
screen "0113_SettingShiftPlan" 1280x800, template "Navigation"
   on GenerateScreen: SetTag("Recipe_Appearance_Control", 1); function_b431313b("Shifttime", U 1, N)
   on ClearScreen: function_f38ba6b2("Shifttime", U 1, 1, 0, N)
   Button "Button_1" at 612,704 size 245x55; TextOff 'Next Shift'
   TextField "Text field_8" at 305,167 size 204x48; Text 'Shift 1'
   TextField "Text field_9" at 517,167 size 204x48; Text 'Shift 2'
   TextField "Text field_10" at 729,167 size 204x48; Text 'Shift 3'
   TextField "Text field_11" at 941,167 size 204x48; Text 'Shift 4'
   Button "Button_3" at 326,104 size 451x32; TextOff 'Setting Shift Plan'
   Button "b_ShifProto_ShotCounter_1" at 208,713 size 60x60; TextOff 'Shot Counter'; PictureList "ico_ShiftProtocol"
      Appearance <- "Recipe_Appearance_Control"
      ProcessValue <- "Recipe_Appearance_Control"
   Button "b_Shiftproto_shiftproto" at 208,713 size 60x60; TextOff 'Shift proto'
      Appearance <- "Recipe_Appearance_Control"
      on Click: ActivateScreen("0112_Shift protocol", 0); SetTag("Recipe_Appearance_Control", 2)
   Button "b_SC" at 478,713 size 60x60; TextOff 'Shot Counter'; PictureList "ico_ShotCounter"
      on Press: ActivateScreen("0891_Shotcounter MixingHead", 0); SetTag("Recipe_Appearance_Control", 5)
      Appearance <- "Recipe_Appearance_Control"
      ProcessValue <- "Recipe_Appearance_Control"
   Button "b_SC_1" at 478,713 size 60x60; TextOff 'Shot Counter'
      Appearance <- "Recipe_Appearance_Control"
      on Click: ActivateScreen("0891_Shotcounter MixingHead", 0); SetTag("Recipe_Appearance_Control", 5)
   Button "b_Shift_Plan" at 118,713 size 60x60; TextOff 'Shift Plan'; PictureList "ico_ShiftPlan"
      on Press: ActivateScreen("0113_SettingShiftPlan", 0); SetTag("Recipe_Appearance_Control", 1)
      Appearance <- "Recipe_Appearance_Control"
      ProcessValue <- "Recipe_Appearance_Control"
   Button "b_Shift_Plan_1" at 118,713 size 60x60; TextOff 'Shift Plan'
      Appearance <- "Recipe_Appearance_Control"
      on Click: "SettingShiftPlan"(); ActivateScreen("0113_SettingShiftPlan", 0); SetTag("Recipe_Appearance_Control", 1)
   Button "b_LS_Lastshot" at 298,713 size 60x60; TextOff 'Last Shot'; PictureList "ico_LastShot"
      on Press: ActivateScreen("0036_Last Shot", 0); SetTag("Recipe_Appearance_Control", 3)
      Appearance <- "Recipe_Appearance_Control"
      ProcessValue <- "Recipe_Appearance_Control"
   Button "b_LS_Lastshot_1" at 298,713 size 60x60; TextOff 'Last Shot'
      Appearance <- "Recipe_Appearance_Control"
      on Click: ActivateScreen("0036_Last Shot", 0); SetTag("Recipe_Appearance_Control", 3)
   Button "b_Consumtion" at 388,713 size 60x60; TextOff 'Consumtion / Consum'; PictureList "ico_consum"
      on Press: ActivateScreen("0890_Consumption", 0); SetTag("Recipe_Appearance_Control", 4)
      Appearance <- "Recipe_Appearance_Control"
      ProcessValue <- "Recipe_Appearance_Control"
   Button "b_Consumtion_1" at 388,713 size 60x60; TextOff 'Consumtion / Consum'
      Appearance <- "Recipe_Appearance_Control"
      on Click: ActivateScreen("0890_Consumption", 0); SetTag("Recipe_Appearance_Control", 4)
   TextField "Text field_1" at 134,234 size 152x60; Text 'Monday'
   TextField "Text field_2" at 134,298 size 152x60; Text 'Tuesday'
   TextField "Text field_3" at 134,362 size 152x60; Text 'Wenesday'
   TextField "Text field_4" at 134,426 size 152x60; Text 'Thrusday'
   TextField "Text field_5" at 134,490 size 152x60; Text 'Friday'
   TextField "Text field_6" at 134,554 size 152x60; Text 'Saturday'
   TextField "Text field_7" at 134,618 size 152x60; Text 'Sunday'
   IOField "I/O field_1" at 303,298 size 135x60; Authorization "Operate"; FormatPattern 9999999999999999999999999999999999999999
      on OnFinishInput: "SettingShiftPlan"(); "Shifttime_write"()
      ProcessValue <- "Shift_2_1"
   IOField "I/O field_2" at 303,362 size 135x60; Authorization "Operate"; FormatPattern 9999999999999999999999999999999999999999
      on OnFinishInput: "SettingShiftPlan"(); "Shifttime_write"()
      ProcessValue <- "Shift_3_1"
   IOField "I/O field_3" at 303,426 size 135x60; Authorization "Operate"; FormatPattern 9999999999999999999999999999999999999999
      on OnFinishInput: "SettingShiftPlan"(); "Shifttime_write"()
      ProcessValue <- "Shift_4_1"
   IOField "I/O field_4" at 303,490 size 135x60; Authorization "Operate"; FormatPattern 9999999999999999999999999999999999999999
      on OnFinishInput: "SettingShiftPlan"(); "Shifttime_write"()
      ProcessValue <- "Shift_5_1"
   IOField "I/O field_5" at 303,554 size 135x60; Authorization "Operate"; FormatPattern 9999999999999999999999999999999999999999
      on OnFinishInput: "SettingShiftPlan"(); "Shifttime_write"()
      ProcessValue <- "Shift_6_1"
   IOField "I/O field_6" at 303,618 size 135x60; Authorization "Operate"; FormatPattern 9999999999999999999999999999999999999999
      on OnFinishInput: "SettingShiftPlan"(); "Shifttime_write"()
      ProcessValue <- "Shift_7_1"
   IOField "I/O field_7" at 303,234 size 135x60; Authorization "Operate"; FormatPattern 9999999999999999999999999999999999999999
      on OnFinishInput: "SettingShiftPlan"(); "Shifttime_write"()
      ProcessValue <- "Shift_1_1"
   IOField "I/O field_8" at 515,298 size 135x60; Authorization "Operate"; FormatPattern 9999999999999999999999999999999999999999
      on OnFinishInput: "SettingShiftPlan"(); "Shifttime_write"()
      ProcessValue <- "Shift_2_2"
   IOField "I/O field_9" at 515,362 size 135x60; Authorization "Operate"; FormatPattern 9999999999999999999999999999999999999999
      on OnFinishInput: "SettingShiftPlan"(); "Shifttime_write"()
      ProcessValue <- "Shift_3_2"
   IOField "I/O field_10" at 515,426 size 135x60; Authorization "Operate"; FormatPattern 9999999999999999999999999999999999999999
      on OnFinishInput: "SettingShiftPlan"(); "Shifttime_write"()
      ProcessValue <- "Shift_4_2"
   IOField "I/O field_11" at 515,490 size 135x60; Authorization "Operate"; FormatPattern 9999999999999999999999999999999999999999
      on OnFinishInput: "SettingShiftPlan"(); "Shifttime_write"()
      ProcessValue <- "Shift_5_2"
   IOField "I/O field_12" at 515,554 size 135x60; Authorization "Operate"; FormatPattern 9999999999999999999999999999999999999999
      on OnFinishInput: "SettingShiftPlan"(); "Shifttime_write"()
      ProcessValue <- "Shift_6_2"
   IOField "I/O field_13" at 515,618 size 135x60; Authorization "Operate"; FormatPattern 9999999999999999999999999999999999999999
      on OnFinishInput: "SettingShiftPlan"(); "Shifttime_write"()
      ProcessValue <- "Shift_7_2"
   IOField "I/O field_14" at 515,234 size 135x60; Authorization "Operate"; FormatPattern 9999999999999999999999999999999999999999
      on OnFinishInput: "SettingShiftPlan"(); "Shifttime_write"()
      ProcessValue <- "Shift_1_2"
   IOField "I/O field_15" at 727,298 size 135x60; Authorization "Operate"; FormatPattern 9999999999999999999999999999999999999999
      on OnFinishInput: "SettingShiftPlan"(); "Shifttime_write"()
      ProcessValue <- "Shift_2_3"
   IOField "I/O field_16" at 727,362 size 135x60; Authorization "Operate"; FormatPattern 9999999999999999999999999999999999999999
      on OnFinishInput: "SettingShiftPlan"(); "Shifttime_write"()
      ProcessValue <- "Shift_3_3"
   IOField "I/O field_17" at 727,426 size 135x60; Authorization "Operate"; FormatPattern 9999999999999999999999999999999999999999
      on OnFinishInput: "SettingShiftPlan"(); "Shifttime_write"()
      ProcessValue <- "Shift_4_3"
   IOField "I/O field_18" at 727,490 size 135x60; Authorization "Operate"; FormatPattern 9999999999999999999999999999999999999999
      on OnFinishInput: "SettingShiftPlan"(); "Shifttime_write"()
      ProcessValue <- "Shift_5_3"
   IOField "I/O field_19" at 727,554 size 135x60; Authorization "Operate"; FormatPattern 9999999999999999999999999999999999999999
      on OnFinishInput: "SettingShiftPlan"(); "Shifttime_write"()
      ProcessValue <- "Shift_6_3"
   IOField "I/O field_20" at 727,618 size 135x60; Authorization "Operate"; FormatPattern 9999999999999999999999999999999999999999
      on OnFinishInput: "SettingShiftPlan"(); "Shifttime_write"()
      ProcessValue <- "Shift_7_3"
   IOField "I/O field_21" at 727,234 size 135x60; Authorization "Operate"; FormatPattern 9999999999999999999999999999999999999999
      on OnFinishInput: "SettingShiftPlan"(); "Shifttime_write"()
      ProcessValue <- "Shift_1_3"
   IOField "I/O field_23" at 939,298 size 135x60; Authorization "Operate"; FormatPattern 9999999999999999999999999999999999999999
      on OnFinishInput: "SettingShiftPlan"(); "Shifttime_write"()
      ProcessValue <- "Shift_2_4"
   IOField "I/O field_24" at 939,362 size 135x60; Authorization "Operate"; FormatPattern 9999999999999999999999999999999999999999
      on OnFinishInput: "SettingShiftPlan"(); "Shifttime_write"()
      ProcessValue <- "Shift_3_4"
   IOField "I/O field_25" at 939,426 size 135x60; Authorization "Operate"; FormatPattern 9999999999999999999999999999999999999999
      on OnFinishInput: "SettingShiftPlan"(); "Shifttime_write"()
      ProcessValue <- "Shift_4_4"
   IOField "I/O field_26" at 939,490 size 135x60; Authorization "Operate"; FormatPattern 9999999999999999999999999999999999999999
      on OnFinishInput: "SettingShiftPlan"(); "Shifttime_write"()
      ProcessValue <- "Shift_5_4"
   IOField "I/O field_27" at 939,554 size 135x60; Authorization "Operate"; FormatPattern 9999999999999999999999999999999999999999
      on OnFinishInput: "SettingShiftPlan"(); "Shifttime_write"()
      ProcessValue <- "Shift_6_4"
   IOField "I/O field_28" at 939,618 size 135x60; Authorization "Operate"; FormatPattern 9999999999999999999999999999999999999999
      on OnFinishInput: "SettingShiftPlan"(); "Shifttime_write"()
      ProcessValue <- "Shift_7_4"
   IOField "I/O field_29" at 939,234 size 135x60; Authorization "Operate"; FormatPattern 9999999999999999999999999999999999999999
      on OnFinishInput: "SettingShiftPlan"(); "Shifttime_write"()
      ProcessValue <- "Shift_1_4"
   Button "check_shift1_1" at 446,298 size 61x60; TextOff 'Text'; PictureOff "download"; PictureList "Check_Uncheck"; Authorization "Operate"
      on Click: InvertBit("Shift_En_2_1")
      on Change: "SettingShiftPlan"(); "Shifttime_write"()
      ProcessValue <- "Shift_En_2_1"
   Button "check_shift1_2" at 446,362 size 61x60; TextOff 'Text'; PictureOff "download"; PictureList "Check_Uncheck"; Authorization "Operate"
      on Click: InvertBit("Shift_En_3_1")
      on Change: "SettingShiftPlan"(); "Shifttime_write"()
      ProcessValue <- "Shift_En_3_1"
   Button "check_shift1_3" at 446,426 size 61x60; TextOff 'Text'; PictureOff "download"; PictureList "Check_Uncheck"; Authorization "Operate"
      on Click: InvertBit("Shift_En_4_1")
      on Change: "SettingShiftPlan"(); "Shifttime_write"()
      ProcessValue <- "Shift_En_4_1"
   Button "check_shift1_4" at 446,490 size 61x60; TextOff 'Text'; PictureOff "download"; PictureList "Check_Uncheck"; Authorization "Operate"
      on Click: InvertBit("Shift_En_5_1")
      on Change: "SettingShiftPlan"(); "Shifttime_write"()
      ProcessValue <- "Shift_En_5_1"
   Button "check_shift1_5" at 446,554 size 61x60; TextOff 'Text'; PictureOff "download"; PictureList "Check_Uncheck"; Authorization "Operate"
      on Click: InvertBit("Shift_En_6_1")
      on Change: "SettingShiftPlan"(); "Shifttime_write"()
      ProcessValue <- "Shift_En_6_1"
   Button "check_shift1_6" at 446,618 size 61x60; TextOff 'Text'; PictureOff "download"; PictureList "Check_Uncheck"; Authorization "Operate"
      on Click: InvertBit("Shift_En_7_1")
      on Change: "SettingShiftPlan"(); "Shifttime_write"()
      ProcessValue <- "Shift_En_7_1"
   Button "check_shift1_7" at 446,234 size 61x60; TextOff 'Text'; PictureOff "download"; PictureList "Check_Uncheck"; Authorization "Operate"
      on Click: InvertBit("Shift_En_1_1")
      on Change: "SettingShiftPlan"(); "Shifttime_write"()
      ProcessValue <- "Shift_En_1_1"
   Button "check_shift4_1" at 1084,298 size 61x60; TextOff 'Text'; PictureOff "download"; PictureList "Check_Uncheck"; Authorization "Operate"
      on Click: InvertBit("Shift_En_2_4")
      on Change: "SettingShiftPlan"(); "Shifttime_write"()
      ProcessValue <- "Shift_En_2_4"
   Button "check_shift4_2" at 1084,362 size 61x60; TextOff 'Text'; PictureOff "download"; PictureList "Check_Uncheck"; Authorization "Operate"
      on Click: InvertBit("Shift_En_3_4")
      on Change: "SettingShiftPlan"(); "Shifttime_write"()
      ProcessValue <- "Shift_En_3_4"
   Button "check_shift4_3" at 1084,426 size 61x60; TextOff 'Text'; PictureOff "download"; PictureList "Check_Uncheck"; Authorization "Operate"
      on Click: InvertBit("Shift_En_4_4")
      on Change: "SettingShiftPlan"(); "Shifttime_write"()
      ProcessValue <- "Shift_En_4_4"
   Button "check_shift4_4" at 1084,490 size 61x60; TextOff 'Text'; PictureOff "download"; PictureList "Check_Uncheck"; Authorization "Operate"
      on Click: InvertBit("Shift_En_5_4")
      on Change: "SettingShiftPlan"(); "Shifttime_write"()
      ProcessValue <- "Shift_En_5_4"
   Button "check_shift4_5" at 1084,554 size 61x60; TextOff 'Text'; PictureOff "download"; PictureList "Check_Uncheck"; Authorization "Operate"
      on Click: InvertBit("Shift_En_6_4")
      on Change: "SettingShiftPlan"(); "Shifttime_write"()
      ProcessValue <- "Shift_En_6_4"
   Button "check_shift4_6" at 1084,618 size 61x60; TextOff 'Text'; PictureOff "download"; PictureList "Check_Uncheck"; Authorization "Operate"
      on Click: InvertBit("Shift_En_7_4")
      on Change: "SettingShiftPlan"(); "Shifttime_write"()
      ProcessValue <- "Shift_En_7_4"
   Button "check_shift4_7" at 1084,234 size 61x60; TextOff 'Text'; PictureOff "download"; PictureList "Check_Uncheck"; Authorization "Operate"
      on Click: InvertBit("Shift_En_1_4")
      on Change: "SettingShiftPlan"(); "Shifttime_write"()
      ProcessValue <- "Shift_En_1_4"
   Button "check_shift3_1" at 870,298 size 61x60; TextOff 'Text'; PictureOff "download"; PictureList "Check_Uncheck"; Authorization "Operate"
      on Click: InvertBit("Shift_En_2_3")
      on Change: "SettingShiftPlan"(); "Shifttime_write"()
      ProcessValue <- "Shift_En_2_3"
   Button "check_shift3_2" at 870,362 size 61x60; TextOff 'Text'; PictureOff "download"; PictureList "Check_Uncheck"; Authorization "Operate"
      on Click: InvertBit("Shift_En_3_3")
      on Change: "SettingShiftPlan"(); "Shifttime_write"()
      ProcessValue <- "Shift_En_3_3"
   Button "check_shift3_3" at 870,426 size 61x60; TextOff 'Text'; PictureOff "download"; PictureList "Check_Uncheck"; Authorization "Operate"
      on Click: InvertBit("Shift_En_4_3")
      on Change: "SettingShiftPlan"(); "Shifttime_write"()
      ProcessValue <- "Shift_En_4_3"
   Button "check_shift3_4" at 870,490 size 61x60; TextOff 'Text'; PictureOff "download"; PictureList "Check_Uncheck"; Authorization "Operate"
      on Click: InvertBit("Shift_En_5_3")
      on Change: "SettingShiftPlan"(); "Shifttime_write"()
      ProcessValue <- "Shift_En_5_3"
   Button "check_shift3_5" at 870,554 size 61x60; TextOff 'Text'; PictureOff "download"; PictureList "Check_Uncheck"; Authorization "Operate"
      on Click: InvertBit("Shift_En_6_3")
      on Change: "SettingShiftPlan"(); "Shifttime_write"()
      ProcessValue <- "Shift_En_6_3"
   Button "check_shift3_6" at 870,618 size 61x60; TextOff 'Text'; PictureOff "download"; PictureList "Check_Uncheck"; Authorization "Operate"
      on Click: InvertBit("Shift_En_7_3")
      on Change: "SettingShiftPlan"(); "Shifttime_write"()
      ProcessValue <- "Shift_En_7_3"
   Button "check_shift3_7" at 870,234 size 61x60; TextOff 'Text'; PictureOff "download"; PictureList "Check_Uncheck"; Authorization "Operate"
      on Click: InvertBit("Shift_En_1_3")
      on Change: "SettingShiftPlan"(); "Shifttime_write"()
      ProcessValue <- "Shift_En_1_3"
   Button "check_shift2_1" at 659,298 size 61x60; TextOff 'Text'; PictureOff "download"; PictureList "Check_Uncheck"; Authorization "Operate"
      on Click: InvertBit("Shift_En_2_2")
      on Change: "SettingShiftPlan"(); "Shifttime_write"()
      ProcessValue <- "Shift_En_2_2"
   Button "check_shift2_2" at 659,362 size 61x60; TextOff 'Text'; PictureOff "download"; PictureList "Check_Uncheck"; Authorization "Operate"
      on Click: InvertBit("Shift_En_3_2")
      on Change: "SettingShiftPlan"(); "Shifttime_write"()
      ProcessValue <- "Shift_En_3_2"
   Button "check_shift2_3" at 659,426 size 61x60; TextOff 'Text'; PictureOff "download"; PictureList "Check_Uncheck"; Authorization "Operate"
      on Click: InvertBit("Shift_En_4_2")
      on Change: "SettingShiftPlan"(); "Shifttime_write"()
      ProcessValue <- "Shift_En_4_2"
   Button "check_shift2_4" at 659,490 size 61x60; TextOff 'Text'; PictureOff "download"; PictureList "Check_Uncheck"; Authorization "Operate"
      on Click: InvertBit("Shift_En_5_2")
      on Change: "SettingShiftPlan"(); "Shifttime_write"()
      ProcessValue <- "Shift_En_5_2"
   Button "check_shift2_5" at 659,554 size 61x60; TextOff 'Text'; PictureOff "download"; PictureList "Check_Uncheck"; Authorization "Operate"
      on Click: InvertBit("Shift_En_6_2")
      on Change: "SettingShiftPlan"(); "Shifttime_write"()
      ProcessValue <- "Shift_En_6_2"
   Button "check_shift2_6" at 659,618 size 61x60; TextOff 'Text'; PictureOff "download"; PictureList "Check_Uncheck"; Authorization "Operate"
      on Click: InvertBit("Shift_En_7_2")
      on Change: "SettingShiftPlan"(); "Shifttime_write"()
      ProcessValue <- "Shift_En_7_2"
   Button "check_shift2_7" at 659,234 size 61x60; TextOff 'Text'; PictureOff "download"; PictureList "Check_Uncheck"; Authorization "Operate"
      on Click: InvertBit("Shift_En_1_2")
      on Change: "SettingShiftPlan"(); "Shifttime_write"()
      ProcessValue <- "Shift_En_1_2"
   IOField "I/O field_30" at 894,704 size 227x55; FormatPattern 9999999999999999999999999999999999999999
      ProcessValue <- "Next shift"

screen "0112_Shift protocol" 1280x800, template "Navigation"
   on GenerateScreen: SetTag("Recipe_Appearance_Control", 2); function_b431313b("ShiftProtocol", U 1, N)
   on ClearScreen: SetTag("Recipe_Appearance_Control", 0)
   TextField "Text field_1" at 109,205 size 57x47; Text '1.'
   TextField "Text field_2" at 109,270 size 57x47; Text '2.'
   TextField "Text field_3" at 109,335 size 57x47; Text '3.'
   TextField "Text field_4" at 109,402 size 57x47; Text '4.'
   TextField "Text field_5" at 109,469 size 57x47; Text '5.'
   TextField "Text field_6" at 109,537 size 57x47; Text '6.'
   TextField "Text field_7" at 109,605 size 57x47; Text '7.'
   IOField "shiftproto_1" at 176,205 size 267x47; FormatPattern 9999999999999999999999999999999999999999
      ProcessValue <- "Shift_Protocol_1"
   IOField "I/O field_2" at 176,270 size 267x47; FormatPattern 9999999999999999999999999999999999999999
      ProcessValue <- "Shift_Protocol_2"
   IOField "I/O field_3" at 176,335 size 267x47; FormatPattern 9999999999999999999999999999999999999999
      ProcessValue <- "Shift_Protocol_3"
   IOField "I/O field_4" at 176,402 size 267x47; FormatPattern 9999999999999999999999999999999999999999
      ProcessValue <- "Shift_Protocol_4"
   IOField "I/O field_5" at 176,469 size 267x47; FormatPattern 9999999999999999999999999999999999999999
      ProcessValue <- "Shift_Protocol_5"
   IOField "I/O field_6" at 176,537 size 267x47; FormatPattern 9999999999999999999999999999999999999999
      ProcessValue <- "Shift_Protocol_6"
   IOField "I/O field_7" at 176,605 size 267x47; FormatPattern 9999999999999999999999999999999999999999
      ProcessValue <- "Shift_Protocol_7"
   IOField "I/O field_8" at 543,205 size 267x47; FormatPattern 9999999999999999999999999999999999999999
      ProcessValue <- "Shift_Protocol_8"
   IOField "I/O field_9" at 902,205 size 267x47; FormatPattern 9999999999999999999999999999999999999999
      ProcessValue <- "Shift_Protocol_15"
   IOField "I/O field_10" at 543,270 size 267x47; FormatPattern 9999999999999999999999999999999999999999
      ProcessValue <- "Shift_Protocol_9"
   IOField "I/O field_11" at 543,335 size 267x47; FormatPattern 9999999999999999999999999999999999999999
      ProcessValue <- "Shift_Protocol_10"
   IOField "I/O field_12" at 543,402 size 267x47; FormatPattern 9999999999999999999999999999999999999999
      ProcessValue <- "Shift_Protocol_11"
   IOField "I/O field_13" at 543,469 size 267x47; FormatPattern 9999999999999999999999999999999999999999
      ProcessValue <- "Shift_Protocol_12"
   IOField "I/O field_14" at 543,537 size 267x47; FormatPattern 9999999999999999999999999999999999999999
      ProcessValue <- "Shift_Protocol_13"
   IOField "I/O field_15" at 543,605 size 267x47; FormatPattern 9999999999999999999999999999999999999999
      ProcessValue <- "Shift_Protocol_14"
   IOField "I/O field_16" at 902,270 size 267x47; FormatPattern 9999999999999999999999999999999999999999
      ProcessValue <- "Shift_Protocol_16"
   IOField "I/O field_17" at 902,335 size 267x47; FormatPattern 9999999999999999999999999999999999999999
      ProcessValue <- "Shift_Protocol_17"
   IOField "I/O field_18" at 902,402 size 267x47; FormatPattern 9999999999999999999999999999999999999999
      ProcessValue <- "Shift_Protocol_18"
   IOField "I/O field_19" at 902,469 size 267x47; FormatPattern 9999999999999999999999999999999999999999
      ProcessValue <- "Shift_Protocol_19"
   IOField "I/O field_20" at 902,537 size 267x47; FormatPattern 9999999999999999999999999999999999999999
      ProcessValue <- "Shift_Protocol_20"
   IOField "I/O field_21" at 902,605 size 267x47; FormatPattern 9999999999999999999999999999999999999999
      ProcessValue <- "Shift_Protocol_21"
   TextField "Text field_8" at 474,205 size 57x47; Text '8.'
   TextField "Text field_9" at 474,270 size 57x47; Text '9.'
   TextField "Text field_10" at 474,335 size 57x47; Text '10.'
   TextField "Text field_11" at 474,402 size 57x47; Text '11.'
   TextField "Text field_12" at 474,469 size 57x47; Text '12.'
   TextField "Text field_13" at 474,537 size 57x47; Text '13.'
   TextField "Text field_14" at 474,605 size 57x47; Text '14.'
   TextField "Text field_15" at 836,205 size 57x47; Text '15.'
   TextField "Text field_16" at 836,270 size 57x47; Text '16.'
   TextField "Text field_17" at 836,335 size 57x47; Text '17.'
   TextField "Text field_18" at 836,402 size 57x47; Text '18.'
   TextField "Text field_19" at 836,469 size 57x47; Text '19.'
   TextField "Text field_20" at 836,537 size 57x47; Text '20.'
   TextField "Text field_21" at 836,605 size 57x47; Text '21.'
   Button "Button_3" at 326,104 size 451x32; TextOff 'Shift Protocol'
   Button "b_spare" at 1000,713 size 60x60; TextOff 'Text'; PictureOff "USB_1"
      on Click: function_ea909784("ShiftProtocol", U 0, '\Storage Card USB\record.csv', 1, 1, N)
   Button "Button_1" at 172,202 size 276x54; TextOff 'Text'
      on Click: SetTag("Archive Alarm Number", 1); SetTag("Archived Alarm Control", 1); "CopyAlarmLogView"(); ActivateScreen("0013_Archive Alarm", 0)
   Button "b_ShifProto_ShotCounter_1" at 208,713 size 60x60; TextOff 'Shot Counter'; PictureList "ico_ShiftProtocol"
      ProcessValue <- "Recipe_Appearance_Control"
      Appearance <- "Recipe_Appearance_Control"
   Button "b_Shiftproto_shiftproto" at 208,713 size 60x60; TextOff 'Shift proto'
      on Click: ActivateScreen("0112_Shift protocol", 0); SetTag("Recipe_Appearance_Control", 2)
      Appearance <- "Recipe_Appearance_Control"
   Button "b_SC" at 478,713 size 60x60; TextOff 'Shot Counter'; PictureList "ico_ShotCounter"
      on Press: ActivateScreen("0891_Shotcounter MixingHead", 0); SetTag("Recipe_Appearance_Control", 5)
      Appearance <- "Recipe_Appearance_Control"
      ProcessValue <- "Recipe_Appearance_Control"
   Button "b_SC_1" at 478,713 size 60x60; TextOff 'Shot Counter'
      on Click: ActivateScreen("0891_Shotcounter MixingHead", 0); SetTag("Recipe_Appearance_Control", 5)
      Appearance <- "Recipe_Appearance_Control"
   Button "b_Shift_Plan" at 118,713 size 60x60; TextOff 'Shift Plan'; PictureList "ico_ShiftPlan"
      on Press: ActivateScreen("0113_SettingShiftPlan", 0); SetTag("Recipe_Appearance_Control", 1)
      Appearance <- "Recipe_Appearance_Control"
      ProcessValue <- "Recipe_Appearance_Control"
   Button "b_Shift_Plan_1" at 118,713 size 60x60; TextOff 'Shift Plan'
      on Click: "SettingShiftPlan"(); ActivateScreen("0113_SettingShiftPlan", 0); SetTag("Recipe_Appearance_Control", 1)
      Appearance <- "Recipe_Appearance_Control"
   Button "b_LS_Lastshot" at 298,713 size 60x60; TextOff 'Last Shot'; PictureList "ico_LastShot"
      on Press: ActivateScreen("0036_Last Shot", 0); SetTag("Recipe_Appearance_Control", 3)
      Appearance <- "Recipe_Appearance_Control"
      ProcessValue <- "Recipe_Appearance_Control"
   Button "b_LS_Lastshot_1" at 298,713 size 60x60; TextOff 'Last Shot'
      on Click: ActivateScreen("0036_Last Shot", 0); SetTag("Recipe_Appearance_Control", 3)
      Appearance <- "Recipe_Appearance_Control"
   Button "b_Consumtion" at 388,713 size 60x60; TextOff 'Consumtion / Consum'; PictureList "ico_consum"
      on Press: ActivateScreen("0890_Consumption", 0); SetTag("Recipe_Appearance_Control", 4)
      Appearance <- "Recipe_Appearance_Control"
      ProcessValue <- "Recipe_Appearance_Control"
   Button "b_Consumtion_1" at 388,713 size 60x60; TextOff 'Consumtion / Consum'
      on Click: ActivateScreen("0890_Consumption", 0); SetTag("Recipe_Appearance_Control", 4)
      Appearance <- "Recipe_Appearance_Control"
   Button "Button_2" at 172,267 size 276x54; TextOff 'Text'
      on Click: SetTag("Archive Alarm Number", 2); SetTag("Archived Alarm Control", 1); "CopyAlarmLogView"(); ActivateScreen("0013_Archive Alarm", 0)
   Button "Button_4" at 172,332 size 276x54; TextOff 'Text'
      on Click: SetTag("Archive Alarm Number", 3); SetTag("Archived Alarm Control", 1); "CopyAlarmLogView"(); ActivateScreen("0013_Archive Alarm", 0)
   Button "Button_5" at 172,397 size 276x54; TextOff 'Text'
      on Click: SetTag("Archive Alarm Number", 4); SetTag("Archived Alarm Control", 1); "CopyAlarmLogView"(); ActivateScreen("0013_Archive Alarm", 0)
   Button "Button_6" at 172,465 size 276x54; TextOff 'Text'
      on Click: SetTag("Archive Alarm Number", 5); SetTag("Archived Alarm Control", 1); "CopyAlarmLogView"(); ActivateScreen("0013_Archive Alarm", 0)
   Button "Button_7" at 172,535 size 276x54; TextOff 'Text'
      on Click: SetTag("Archive Alarm Number", 6); SetTag("Archived Alarm Control", 1); "CopyAlarmLogView"(); ActivateScreen("0013_Archive Alarm", 0)
   Button "Button_8" at 172,602 size 276x54; TextOff 'Text'
      on Click: SetTag("Archive Alarm Number", 7); SetTag("Archived Alarm Control", 1); "CopyAlarmLogView"(); ActivateScreen("0013_Archive Alarm", 0)
   Button "Button_9" at 540,202 size 276x54; TextOff 'Text'
      on Click: SetTag("Archive Alarm Number", 8); SetTag("Archived Alarm Control", 1); "CopyAlarmLogView"(); ActivateScreen("0013_Archive Alarm", 0)
   Button "Button_10" at 540,267 size 276x54; TextOff 'Text'
      on Click: SetTag("Archive Alarm Number", 9); SetTag("Archived Alarm Control", 1); "CopyAlarmLogView"(); ActivateScreen("0013_Archive Alarm", 0)
   Button "Button_11" at 540,332 size 276x54; TextOff 'Text'
      on Click: SetTag("Archive Alarm Number", 10); SetTag("Archived Alarm Control", 1); "CopyAlarmLogView"(); ActivateScreen("0013_Archive Alarm", 0)
   Button "Button_12" at 540,397 size 276x54; TextOff 'Text'
      on Click: SetTag("Archive Alarm Number", 11); SetTag("Archived Alarm Control", 1); "CopyAlarmLogView"(); ActivateScreen("0013_Archive Alarm", 0)
   Button "Button_13" at 540,465 size 276x54; TextOff 'Text'
      on Click: SetTag("Archive Alarm Number", 12); SetTag("Archived Alarm Control", 1); "CopyAlarmLogView"(); ActivateScreen("0013_Archive Alarm", 0)
   Button "Button_14" at 540,535 size 276x54; TextOff 'Text'
      on Click: SetTag("Archive Alarm Number", 13); SetTag("Archived Alarm Control", 1); "CopyAlarmLogView"(); ActivateScreen("0013_Archive Alarm", 0)
   Button "Button_15" at 540,602 size 276x54; TextOff 'Text'
      on Click: SetTag("Archive Alarm Number", 14); SetTag("Archived Alarm Control", 1); "CopyAlarmLogView"(); ActivateScreen("0013_Archive Alarm", 0)
   Button "Button_16" at 900,202 size 276x54; TextOff 'Text'
      on Click: SetTag("Archive Alarm Number", 15); SetTag("Archived Alarm Control", 1); "CopyAlarmLogView"(); ActivateScreen("0013_Archive Alarm", 0)
   Button "Button_17" at 900,267 size 276x54; TextOff 'Text'
      on Click: SetTag("Archive Alarm Number", 16); SetTag("Archived Alarm Control", 1); "CopyAlarmLogView"(); ActivateScreen("0013_Archive Alarm", 0)
   Button "Button_18" at 900,332 size 276x54; TextOff 'Text'
      on Click: SetTag("Archive Alarm Number", 17); SetTag("Archived Alarm Control", 1); "CopyAlarmLogView"(); ActivateScreen("0013_Archive Alarm", 0)
   Button "Button_19" at 900,397 size 276x54; TextOff 'Text'
      on Click: SetTag("Archive Alarm Number", 18); SetTag("Archived Alarm Control", 1); "CopyAlarmLogView"(); ActivateScreen("0013_Archive Alarm", 0)
   Button "Button_20" at 900,465 size 276x54; TextOff 'Text'
      on Click: SetTag("Archive Alarm Number", 19); SetTag("Archived Alarm Control", 1); "CopyAlarmLogView"(); ActivateScreen("0013_Archive Alarm", 0)
   Button "Button_21" at 900,535 size 276x54; TextOff 'Text'
      on Click: SetTag("Archive Alarm Number", 20); SetTag("Archived Alarm Control", 1); "CopyAlarmLogView"(); ActivateScreen("0013_Archive Alarm", 0)
   Button "Button_22" at 900,602 size 276x54; TextOff 'Text'
      on Click: SetTag("Archive Alarm Number", 21); SetTag("Archived Alarm Control", 1); "CopyAlarmLogView"(); ActivateScreen("0013_Archive Alarm", 0)

screen "0036_Last Shot" 1280x800, template "Navigation"
   on GenerateScreen: SetTag("Recipe_Appearance_Control", 3)
   IOField "Prg_1" at 156,204 size 45x30; FormatPattern 99
      ProcessValue <- "DB918_ShotResultlast10_FilteredShot{1}_StationNo"
   IOField "I/O field_2" at 156,290 size 45x30; FormatPattern 99
      ProcessValue <- "DB918_ShotResultlast10_FilteredShot{2}_StationNo"
   IOField "I/O field_3" at 156,378 size 45x30; FormatPattern 99
      ProcessValue <- "DB918_ShotResultlast10_FilteredShot{3}_StationNo"
   IOField "I/O field_4" at 156,466 size 45x30; FormatPattern 99
      ProcessValue <- "DB918_ShotResultlast10_FilteredShot{4}_StationNo"
   IOField "I/O field_5" at 156,551 size 45x30; FormatPattern 99
      ProcessValue <- "DB918_ShotResultlast10_FilteredShot{5}_StationNo"
   IOField "I/O field_6" at 156,637 size 45x30; FormatPattern 99
      ProcessValue <- "DB918_ShotResultlast10_FilteredShot{6}_StationNo"
   IOField "I/O field_7" at 209,204 size 45x30; FormatPattern 99
      ProcessValue <- "DB918_ShotResultlast10_FilteredShot{1}_MHNo"
   IOField "I/O field_8" at 209,290 size 45x30; FormatPattern 99
      ProcessValue <- "DB918_ShotResultlast10_FilteredShot{2}_MHNo"
   IOField "I/O field_9" at 209,378 size 45x30; FormatPattern 99
      ProcessValue <- "DB918_ShotResultlast10_FilteredShot{3}_MHNo"
   IOField "I/O field_10" at 209,466 size 45x30; FormatPattern 99
      ProcessValue <- "DB918_ShotResultlast10_FilteredShot{4}_MHNo"
   IOField "I/O field_11" at 209,551 size 45x30; FormatPattern 99
      ProcessValue <- "DB918_ShotResultlast10_FilteredShot{5}_MHNo"
   IOField "I/O field_12" at 209,637 size 45x30; FormatPattern 99
      ProcessValue <- "DB918_ShotResultlast10_FilteredShot{6}_MHNo"
   IOField "I/O field_13" at 262,204 size 45x30; FormatPattern 99
      ProcessValue <- "DB918_ShotResultlast10_FilteredShot{1}_PartNo"
   IOField "I/O field_14" at 262,290 size 45x30; FormatPattern 99
      ProcessValue <- "DB918_ShotResultlast10_FilteredShot{2}_PartNo"
   IOField "I/O field_15" at 262,378 size 45x30; FormatPattern 99
      ProcessValue <- "DB918_ShotResultlast10_FilteredShot{3}_PartNo"
   IOField "I/O field_16" at 262,466 size 45x30; FormatPattern 99
      ProcessValue <- "DB918_ShotResultlast10_FilteredShot{4}_PartNo"
   IOField "I/O field_17" at 262,551 size 45x30; FormatPattern 99
      ProcessValue <- "DB918_ShotResultlast10_FilteredShot{5}_PartNo"
   IOField "I/O field_18" at 262,637 size 45x30; FormatPattern 99
      ProcessValue <- "DB918_ShotResultlast10_FilteredShot{6}_PartNo"
   IOField "I/O field_19" at 314,204 size 102x30; FormatPattern 9999.999
      ProcessValue <- "DB918_ShotResultlast10_FilteredShot{1}_FoamingTime"
   IOField "I/O field_20" at 314,290 size 102x30; FormatPattern 9999.999
      ProcessValue <- "DB918_ShotResultlast10_FilteredShot{2}_FoamingTime"
   IOField "I/O field_21" at 314,378 size 102x30; FormatPattern 9999.999
      ProcessValue <- "DB918_ShotResultlast10_FilteredShot{3}_FoamingTime"
   IOField "I/O field_22" at 314,466 size 102x30; FormatPattern 9999.999
      ProcessValue <- "DB918_ShotResultlast10_FilteredShot{4}_FoamingTime"
   IOField "I/O field_23" at 314,551 size 102x30; FormatPattern 9999.999
      ProcessValue <- "DB918_ShotResultlast10_FilteredShot{5}_FoamingTime"
   IOField "I/O field_24" at 314,637 size 102x30; FormatPattern 9999.999
      ProcessValue <- "DB918_ShotResultlast10_FilteredShot{6}_FoamingTime"
   IOField "I/O field_25" at 422,204 size 102x30; FormatPattern 999999.99
      ProcessValue <- "DB918_ShotResultlast10_FilteredShot{1}_PartWeight"
   IOField "I/O field_26" at 422,290 size 102x30; FormatPattern 999999.99
      ProcessValue <- "DB918_ShotResultlast10_FilteredShot{2}_PartWeight"
   IOField "I/O field_27" at 422,378 size 102x30; FormatPattern 999999.99
      ProcessValue <- "DB918_ShotResultlast10_FilteredShot{3}_PartWeight"
   IOField "I/O field_28" at 422,466 size 102x30; FormatPattern 999999.99
      ProcessValue <- "DB918_ShotResultlast10_FilteredShot{4}_PartWeight"
   IOField "I/O field_29" at 422,551 size 102x30; FormatPattern 999999.99
      ProcessValue <- "DB918_ShotResultlast10_FilteredShot{5}_PartWeight"
   IOField "I/O field_30" at 422,637 size 102x30; FormatPattern 999999.99
      ProcessValue <- "DB918_ShotResultlast10_FilteredShot{6}_PartWeight"
   IOField "I/O field_31" at 717,204 size 102x30; FormatPattern 999999.99
      ProcessValue <- "DB918_ShotResultlast10_FilteredShot{1}_Flow{1}"
   IOField "I/O field_32" at 717,240 size 102x30; FormatPattern 999999.99
      ProcessValue <- "DB918_ShotResultlast10_FilteredShot{1}_Flow{2}"
   IOField "I/O field_33" at 717,290 size 102x30; FormatPattern 999999.99
      ProcessValue <- "DB918_ShotResultlast10_FilteredShot{2}_Flow{1}"
   IOField "I/O field_34" at 717,327 size 102x30; FormatPattern 999999.99
      ProcessValue <- "DB918_ShotResultlast10_FilteredShot{2}_Flow{2}(1)"
   IOField "I/O field_35" at 717,379 size 102x30; FormatPattern 999999.99
      ProcessValue <- "DB918_ShotResultlast10_FilteredShot{3}_Flow{1}"
   IOField "I/O field_36" at 717,413 size 102x30; FormatPattern 999999.99
      ProcessValue <- "DB918_ShotResultlast10_FilteredShot{3}_Flow{2}"
   IOField "I/O field_37" at 717,466 size 102x30; FormatPattern 999999.99
      ProcessValue <- "DB918_ShotResultlast10_FilteredShot{4}_Flow{1}"
   IOField "I/O field_38" at 717,501 size 102x30; FormatPattern 999999.99
      ProcessValue <- "DB918_ShotResultlast10_FilteredShot{4}_Flow{2}"
   IOField "I/O field_39" at 717,551 size 102x30; FormatPattern 999999.99
      ProcessValue <- "DB918_ShotResultlast10_FilteredShot{5}_Flow{1}"
   IOField "I/O field_40" at 717,586 size 102x30; FormatPattern 999999.99
      ProcessValue <- "DB918_ShotResultlast10_FilteredShot{5}_Flow{2}"
   IOField "I/O field_41" at 717,637 size 102x30; FormatPattern 999999.99
      ProcessValue <- "DB918_ShotResultlast10_FilteredShot{6}_Flow{1}"
   IOField "I/O field_42" at 824,204 size 82x30; FormatPattern 999999.99
      ProcessValue <- "DB918_ShotResultlast10_FilteredShot{1}_Pressure{1}"
   IOField "I/O field_43" at 824,240 size 82x30; FormatPattern 999999.99
      ProcessValue <- "DB918_ShotResultlast10_FilteredShot{1}_Pressure{2}"
   IOField "I/O field_44" at 824,290 size 82x30; FormatPattern 999999.99
      ProcessValue <- "DB918_ShotResultlast10_FilteredShot{2}_Pressure{1}"
   IOField "I/O field_45" at 824,327 size 82x30; FormatPattern 999999.99
      ProcessValue <- "DB918_ShotResultlast10_FilteredShot{2}_Pressure{2}"
   IOField "I/O field_46" at 824,378 size 82x30; FormatPattern 999999.99
      ProcessValue <- "DB918_ShotResultlast10_FilteredShot{3}_Pressure{1}"
   IOField "I/O field_47" at 824,413 size 82x30; FormatPattern 999999.99
      ProcessValue <- "DB918_ShotResultlast10_FilteredShot{3}_Pressure{2}"
   IOField "I/O field_48" at 824,466 size 82x30; FormatPattern 999999.99
      ProcessValue <- "DB918_ShotResultlast10_FilteredShot{4}_Pressure{1}"
   IOField "I/O field_49" at 824,501 size 82x30; FormatPattern 999999.99
      ProcessValue <- "DB918_ShotResultlast10_FilteredShot{4}_Pressure{2}"
   IOField "I/O field_50" at 824,551 size 82x30; FormatPattern 999999.99
      ProcessValue <- "DB918_ShotResultlast10_FilteredShot{5}_Pressure{1}"
   IOField "I/O field_51" at 824,586 size 82x30; FormatPattern 999999.99
      ProcessValue <- "DB918_ShotResultlast10_FilteredShot{5}_Pressure{2}"
   IOField "I/O field_52" at 824,637 size 82x30; FormatPattern 999999.99
      ProcessValue <- "DB918_ShotResultlast10_FilteredShot{6}_Pressure{1}"
   IOField "I/O field_53" at 911,204 size 82x30; FormatPattern 999999.99
      ProcessValue <- "DB918_ShotResultlast10_FilteredShot{1}_Mixingratio{1}"
   IOField "I/O field_54" at 911,240 size 82x30; FormatPattern 999999.99
      ProcessValue <- "DB918_ShotResultlast10_FilteredShot{1}_Mixingratio{2}"
   IOField "I/O field_55" at 911,290 size 82x30; FormatPattern 999999.99
      ProcessValue <- "DB918_ShotResultlast10_FilteredShot{2}_Mixingratio{1}"
   IOField "I/O field_56" at 911,327 size 82x30; FormatPattern 999999.99
      ProcessValue <- "DB918_ShotResultlast10_FilteredShot{2}_Mixingratio{2}"
   IOField "I/O field_57" at 911,379 size 82x30; FormatPattern 999999.99
      ProcessValue <- "DB918_ShotResultlast10_FilteredShot{3}_Mixingratio{1}"
   IOField "I/O field_58" at 911,413 size 82x30; FormatPattern 999999.99
      ProcessValue <- "DB918_ShotResultlast10_FilteredShot{3}_Mixingratio{2}"
   IOField "I/O field_59" at 911,466 size 82x30; FormatPattern 999999.99
      ProcessValue <- "DB918_ShotResultlast10_FilteredShot{4}_Mixingratio{1}"
   IOField "I/O field_60" at 911,501 size 82x30; FormatPattern 999999.99
      ProcessValue <- "DB918_ShotResultlast10_FilteredShot{4}_Mixingratio{2}"
   IOField "I/O field_61" at 911,551 size 82x30; FormatPattern 999999.99
      ProcessValue <- "DB918_ShotResultlast10_FilteredShot{5}_Mixingratio{1}"
   IOField "I/O field_62" at 911,586 size 82x30; FormatPattern 999999.99
      ProcessValue <- "DB918_ShotResultlast10_FilteredShot{5}_Mixingratio{2}"
   IOField "I/O field_63" at 911,637 size 82x30; FormatPattern 999999.99
      ProcessValue <- "DB918_ShotResultlast10_FilteredShot{6}_Mixingratio{1}"
   IOField "I/O field_64" at 998,204 size 82x30; FormatPattern 999999.9
      ProcessValue <- "DB918_ShotResultlast10_FilteredShot{1}_Temperature{1}"
   IOField "I/O field_65" at 998,240 size 82x30; FormatPattern 999999.9
      ProcessValue <- "DB918_ShotResultlast10_FilteredShot{1}_Temperature{2}"
   IOField "I/O field_66" at 998,290 size 82x30; FormatPattern 999999.9
      ProcessValue <- "DB918_ShotResultlast10_FilteredShot{2}_Temperature{1}"
   IOField "I/O field_67" at 998,327 size 82x30; FormatPattern 999999.9
      ProcessValue <- "DB918_ShotResultlast10_FilteredShot{2}_Temperature{2}"
   IOField "I/O field_68" at 998,378 size 82x30; FormatPattern 999999.9
      ProcessValue <- "DB918_ShotResultlast10_FilteredShot{3}_Temperature{1}"
   IOField "I/O field_69" at 998,413 size 82x30; FormatPattern 999999.9
      ProcessValue <- "DB918_ShotResultlast10_FilteredShot{3}_Temperature{2}"
   IOField "I/O field_70" at 998,466 size 82x30; FormatPattern 999999.9
      ProcessValue <- "DB918_ShotResultlast10_FilteredShot{4}_Temperature{1}"
   IOField "I/O field_71" at 998,501 size 82x30; FormatPattern 999999.9
      ProcessValue <- "DB918_ShotResultlast10_FilteredShot{4}_Temperature{2}"
   IOField "I/O field_72" at 998,551 size 82x30; FormatPattern 999999.9
      ProcessValue <- "DB918_ShotResultlast10_FilteredShot{5}_Temperature{1}"
   IOField "I/O field_73" at 998,586 size 82x30; FormatPattern 999999.9
      ProcessValue <- "DB918_ShotResultlast10_FilteredShot{5}_Temperature{2}"
   IOField "I/O field_74" at 998,637 size 82x30; FormatPattern 999999.9
      ProcessValue <- "DB918_ShotResultlast10_FilteredShot{6}_Temperature{1}"
   IOField "I/O field_75" at 1085,204 size 82x30; FormatPattern 999999.99
      ProcessValue <- "DB918_ShotResultlast10_FilteredShot{1}_MaterialConsumption{1}"
   IOField "I/O field_76" at 1085,240 size 82x30; FormatPattern 999999.99
      ProcessValue <- "DB918_ShotResultlast10_FilteredShot{1}_MaterialConsumption{2}"
   IOField "I/O field_77" at 1085,290 size 82x30; FormatPattern 999999.99
      ProcessValue <- "DB918_ShotResultlast10_FilteredShot{2}_MaterialConsumption{1}"
   IOField "I/O field_78" at 1085,327 size 82x30; FormatPattern 999999.99
      ProcessValue <- "DB918_ShotResultlast10_FilteredShot{2}_MaterialConsumption{2}"
   IOField "I/O field_79" at 1085,378 size 82x30; FormatPattern 999999.99
      ProcessValue <- "DB918_ShotResultlast10_FilteredShot{3}_MaterialConsumption{1}"
   IOField "I/O field_80" at 1085,413 size 82x30; FormatPattern 999999.99
      ProcessValue <- "DB918_ShotResultlast10_FilteredShot{3}_MaterialConsumption{2}"
   IOField "I/O field_81" at 1085,466 size 82x30; FormatPattern 999999.99
      ProcessValue <- "DB918_ShotResultlast10_FilteredShot{4}_MaterialConsumption{1}"
   IOField "I/O field_82" at 1085,501 size 82x30; FormatPattern 999999.99
      ProcessValue <- "DB918_ShotResultlast10_FilteredShot{4}_MaterialConsumption{2}"
   IOField "I/O field_83" at 1085,551 size 82x30; FormatPattern 999999.99
      ProcessValue <- "DB918_ShotResultlast10_FilteredShot{5}_MaterialConsumption{1}"
   IOField "I/O field_84" at 1085,586 size 82x30; FormatPattern 999999.99
      ProcessValue <- "DB918_ShotResultlast10_FilteredShot{5}_MaterialConsumption{2}"
   IOField "I/O field_85" at 1085,637 size 82x30; FormatPattern 999999.99
      ProcessValue <- "DB918_ShotResultlast10_FilteredShot{6}_MaterialConsumption{1}"
   Button "Button_3" at 326,99 size 451x32; TextOff 'Last Shot'
   IOField "I/O field_86" at 717,674 size 102x30; FormatPattern 999999.99
      ProcessValue <- "DB918_ShotResultlast10_FilteredShot{6}_Flow{2}"
   IOField "I/O field_87" at 824,674 size 82x30; FormatPattern 999999.99
      ProcessValue <- "DB918_ShotResultlast10_FilteredShot{6}_Pressure{2}"
   IOField "I/O field_88" at 911,674 size 82x30; FormatPattern 999999.99
      ProcessValue <- "DB918_ShotResultlast10_FilteredShot{6}_Mixingratio{2}"
   IOField "I/O field_89" at 998,674 size 82x30; FormatPattern 999999.9
      ProcessValue <- "DB918_ShotResultlast10_FilteredShot{6}_Temperature{2}"
   IOField "I/O field_90" at 1085,674 size 82x30; FormatPattern 999999.99
      ProcessValue <- "DB918_ShotResultlast10_FilteredShot{6}_MaterialConsumption{2}"
   Button "Button_14" at 156,145 size 45x33; TextOff 'Prg.'
   Button "Button_15" at 209,145 size 45x33; TextOff 'MH'
   Button "Button_16" at 262,145 size 45x33; TextOff 'PS'
   Button "Button_17" at 314,145 size 102x33; TextOff 'Time'
   Button "Button_18" at 422,145 size 102x33; TextOff 'Weight'
   Button "Button_19" at 530,145 size 182x33; TextOff 'Name'
   Button "Button_20" at 717,145 size 102x33; TextOff 'Flow'
   Button "Button_21" at 825,145 size 82x33; TextOff 'Pressure'
   Button "Button_22" at 912,145 size 82x33; TextOff 'Ratio'
   Button "Button_23" at 998,145 size 82x33; TextOff 'Temp'
   Button "Button_24" at 1085,145 size 82x33; TextOff 'Weight'
   IOField "I/O field_91" at 529,204 size 182x30; FormatPattern ????????????????????
      ProcessValue <- "DB918_ShotResultlast10_FilteredShot{1}_Name{1}"
   IOField "I/O field_92" at 530,240 size 182x30; FormatPattern ????????????????????
      ProcessValue <- "DB918_ShotResultlast10_FilteredShot{1}_Name{2}"
   IOField "I/O field_93" at 530,290 size 182x30; FormatPattern ????????????????????
      ProcessValue <- "DB918_ShotResultlast10_FilteredShot{2}_Name{1}"
   IOField "I/O field_94" at 530,327 size 182x30; FormatPattern ????????????????????
      ProcessValue <- "DB918_ShotResultlast10_FilteredShot{2}_Name{2}"
   IOField "I/O field_95" at 530,378 size 182x30; FormatPattern ????????????????????
      ProcessValue <- "DB918_ShotResultlast10_FilteredShot{3}_Name{1}"
   IOField "I/O field_96" at 530,413 size 182x30; FormatPattern ????????????????????
      ProcessValue <- "DB918_ShotResultlast10_FilteredShot{3}_Name{2}"
   IOField "I/O field_97" at 530,466 size 182x30; FormatPattern ????????????????????
      ProcessValue <- "DB918_ShotResultlast10_FilteredShot{4}_Name{1}"
   IOField "I/O field_98" at 530,501 size 182x30; FormatPattern ????????????????????
      ProcessValue <- "DB918_ShotResultlast10_FilteredShot{4}_Name{2}"
   IOField "I/O field_99" at 530,551 size 182x30; FormatPattern ????????????????????
      ProcessValue <- "DB918_ShotResultlast10_FilteredShot{5}_Name{1}"
   IOField "I/O field_100" at 530,586 size 182x30; FormatPattern ????????????????????
      ProcessValue <- "DB918_ShotResultlast10_FilteredShot{5}_Name{2}"
   IOField "I/O field_101" at 530,637 size 182x30; FormatPattern ????????????????????
      ProcessValue <- "DB918_ShotResultlast10_FilteredShot{6}_Name{1}"
   IOField "I/O field_102" at 530,674 size 182x30; FormatPattern ????????????????????
      ProcessValue <- "DB918_ShotResultlast10_FilteredShot{6}_Name{2}"
   GraphicView "Graphic view_1" at 104,204 size 45x30; Picture "cp2"
      Visibility <- "DB918_ShotResultlast10_FilteredShot{1}_PartShotDisableService"
   GraphicView "Graphic view_2" at 104,204 size 45x30; Picture "manual mode"
      Visibility <- "DB918_ShotResultlast10_FilteredShot{1}_StatusBitManualShot"
   GraphicView "Graphic view_3" at 104,204 size 45x30; Picture "automatic mode"
      Visibility <- "DB918_ShotResultlast10_FilteredShot{1}_StatusBitAutomaticShot"
   GraphicView "Graphic view_4" at 104,290 size 45x30; Picture "cp2"
      Visibility <- "DB918_ShotResultlast10_FilteredShot{2}_PartShotDisableService"
   GraphicView "Graphic view_5" at 104,290 size 45x30; Picture "manual mode"
      Visibility <- "DB918_ShotResultlast10_FilteredShot{2}_StatusBitManualShot"
   GraphicView "Graphic view_6" at 104,290 size 45x30; Picture "automatic mode"
      Visibility <- "DB918_ShotResultlast10_FilteredShot{2}_StatusBitAutomaticShot"
   GraphicView "Graphic view_7" at 104,378 size 45x30; Picture "cp2"
      Visibility <- "DB918_ShotResultlast10_FilteredShot{3}_PartShotDisableService"
   GraphicView "Graphic view_8" at 104,378 size 45x30; Picture "manual mode"
      Visibility <- "DB918_ShotResultlast10_FilteredShot{3}_StatusBitManualShot"
   GraphicView "Graphic view_9" at 104,378 size 45x30; Picture "automatic mode"
      Visibility <- "DB918_ShotResultlast10_FilteredShot{3}_StatusBitAutomaticShot"
   GraphicView "Graphic view_10" at 104,462 size 45x30; Picture "cp2"
      Visibility <- "DB918_ShotResultlast10_FilteredShot{4}_PartShotDisableService"
   GraphicView "Graphic view_11" at 104,462 size 45x30; Picture "manual mode"
      Visibility <- "DB918_ShotResultlast10_FilteredShot{4}_StatusBitManualShot"
   GraphicView "Graphic view_12" at 104,462 size 45x30; Picture "automatic mode"
      Visibility <- "DB918_ShotResultlast10_FilteredShot{4}_StatusBitAutomaticShot"
   GraphicView "Graphic view_13" at 104,551 size 45x30; Picture "cp2"
      Visibility <- "DB918_ShotResultlast10_FilteredShot{5}_PartShotDisableService"
   GraphicView "Graphic view_14" at 104,551 size 45x30; Picture "manual mode"
      Visibility <- "DB918_ShotResultlast10_FilteredShot{5}_StatusBitManualShot"
   GraphicView "Graphic view_15" at 104,551 size 45x30; Picture "automatic mode"
      Visibility <- "DB918_ShotResultlast10_FilteredShot{5}_StatusBitAutomaticShot"
   GraphicView "Graphic view_16" at 104,637 size 45x30; Picture "cp2"
      Visibility <- "DB918_ShotResultlast10_FilteredShot{6}_PartShotDisableService"
   GraphicView "Graphic view_17" at 104,637 size 45x30; Picture "manual mode"
      Visibility <- "DB918_ShotResultlast10_FilteredShot{6}_StatusBitManualShot"
   GraphicView "Graphic view_18" at 104,637 size 45x30; Picture "automatic mode"
      Visibility <- "DB918_ShotResultlast10_FilteredShot{6}_StatusBitAutomaticShot"
   Button "b_ShifProto_ShotCounter_1" at 208,713 size 60x60; TextOff 'Shot Counter'; PictureList "ico_ShiftProtocol"
      ProcessValue <- "Recipe_Appearance_Control"
      Appearance <- "Recipe_Appearance_Control"
   Button "b_Shiftproto_shiftproto" at 208,713 size 60x60; TextOff 'Shift proto'
      on Click: ActivateScreen("0112_Shift protocol", 0); SetTag("Recipe_Appearance_Control", 2)
      Appearance <- "Recipe_Appearance_Control"
   Button "b_SC" at 478,713 size 60x60; TextOff 'Shot Counter'; PictureList "ico_ShotCounter"
      on Press: ActivateScreen("0891_Shotcounter MixingHead", 0); SetTag("Recipe_Appearance_Control", 5)
      Appearance <- "Recipe_Appearance_Control"
      ProcessValue <- "Recipe_Appearance_Control"
   Button "b_SC_1" at 478,713 size 60x60; TextOff 'Shot Counter'
      on Click: ActivateScreen("0891_Shotcounter MixingHead", 0); SetTag("Recipe_Appearance_Control", 5)
      Appearance <- "Recipe_Appearance_Control"
   Button "b_Shift_Plan" at 118,713 size 60x60; TextOff 'Shift Plan'; PictureList "ico_ShiftPlan"
      on Press: ActivateScreen("0113_SettingShiftPlan", 0); SetTag("Recipe_Appearance_Control", 1)
      Appearance <- "Recipe_Appearance_Control"
      ProcessValue <- "Recipe_Appearance_Control"
   Button "b_Shift_Plan_1" at 118,713 size 60x60; TextOff 'Shift Plan'
      on Click: "SettingShiftPlan"(); ActivateScreen("0113_SettingShiftPlan", 0); SetTag("Recipe_Appearance_Control", 1)
      Appearance <- "Recipe_Appearance_Control"
   Button "b_LS_Lastshot" at 298,713 size 60x60; TextOff 'Last Shot'; PictureList "ico_LastShot"
      on Press: ActivateScreen("0036_Last Shot", 0); SetTag("Recipe_Appearance_Control", 3)
      Appearance <- "Recipe_Appearance_Control"
      ProcessValue <- "Recipe_Appearance_Control"
   Button "b_LS_Lastshot_1" at 298,713 size 60x60; TextOff 'Last Shot'
      on Click: ActivateScreen("0036_Last Shot", 0); SetTag("Recipe_Appearance_Control", 3)
      Appearance <- "Recipe_Appearance_Control"
   Button "b_Consumtion" at 388,713 size 60x60; TextOff 'Consumtion / Consum'; PictureList "ico_consum"
      on Press: ActivateScreen("0890_Consumption", 0); SetTag("Recipe_Appearance_Control", 4)
      Appearance <- "Recipe_Appearance_Control"
      ProcessValue <- "Recipe_Appearance_Control"
   Button "b_Consumtion_1" at 388,713 size 60x60; TextOff 'Consumtion / Consum'
      on Click: ActivateScreen("0890_Consumption", 0); SetTag("Recipe_Appearance_Control", 4)
      Appearance <- "Recipe_Appearance_Control"

